VAR_GLOBAL   // PLC tag table "SDC_Carrier_TagTable"
   "Carrier_01_Carrier_In_Zone" AT %QW400 : Word;
   "Carrier_01_Carrier_Number_Echo" AT %QW402 : Word;
   "Carrier_01_Carrier_Position_Echo" AT %QD404 : DWord;
   "Carrier_01_Next_Carrier_Number" AT %QW408 : Word;
   "Carrier_01_Next_Stop_Position" AT %QD410 : DWord;
   "Carrier_01_Drive_Command_Speed" AT %QW414 : Word;
   "Carrier_01_Duplicate_Carrier_Number" AT %QW416 : Word;
   "Carrier_01_First_Duplicate_Carrier_Position" AT %QD418 : DWord;
   "Carrier_01_Second_Duplicate_Carrier_Position" AT %QD422 : DWord;
   "Carrier_01_CommandWord" AT %QW426 : Word;
   "Carrier_01_Heartbeat" AT %Q426.0 : Bool;
   "Carrier_01_Drive_Forward_Command" AT %Q426.1 : Bool;
   "Carrier_01_Fault_Reset" AT %Q426.2 : Bool;
   "Carrier_01_At_Command_Position" AT %Q426.3 : Bool;
   "Carrier_01_Duplicate_Carrier_Fault" AT %Q426.4 : Bool;
   "Carrier_01_Motion_On_Fault" AT %Q426.5 : Bool;
   "Carrier_01_Motion_Off_Fault" AT %Q426.6 : Bool;
   "Carrier_01_Carrier_Spacing_Fault" AT %Q426.7 : Bool;
   "Carrier_02_Carrier_In_Zone" AT %QW450 : Word;
   "Carrier_02_Carrier_Number_Echo" AT %QW452 : Word;
   "Carrier_02_Carrier_Position_Echo" AT %QD454 : DWord;
   "Carrier_02_Next_Carrier_Number" AT %QW458 : Word;
   "Carrier_02_Next_Stop_Position" AT %QD460 : DWord;
   "Carrier_02_Drive_Command_Speed" AT %QW464 : Word;
   "Carrier_02_Duplicate_Carrier_Number" AT %QW466 : Word;
   "Carrier_02_First_Duplicate_Carrier_Position" AT %QD468 : DWord;
   "Carrier_02_Second_Duplicate_Carrier_Position" AT %QD472 : DWord;
   "Carrier_02_CommandWord" AT %QW476 : Word;
   "Carrier_02_Heartbeat" AT %Q476.0 : Bool;
   "Carrier_02_Drive_Forward_Command" AT %Q476.1 : Bool;
   "Carrier_02_Fault_Reset" AT %Q476.2 : Bool;
   "Carrier_02_At_Command_Position" AT %Q476.3 : Bool;
   "Carrier_02_Duplicate_Carrier_Fault" AT %Q476.4 : Bool;
   "Carrier_02_Motion_On_Fault" AT %Q476.5 : Bool;
   "Carrier_02_Motion_Off_Fault" AT %Q476.6 : Bool;
   "Carrier_02_Carrier_Spacing_Fault" AT %Q476.7 : Bool;
   "Carrier_03_Carrier_In_Zone" AT %QW500 : Word;
   "Carrier_03_Carrier_Number_Echo" AT %QW502 : Word;
   "Carrier_03_Carrier_Position_Echo" AT %QD504 : DWord;
   "Carrier_03_Next_Carrier_Number" AT %QW508 : Word;
   "Carrier_03_Next_Stop_Position" AT %QD510 : DWord;
   "Carrier_03_Drive_Command_Speed" AT %QW514 : Word;
   "Carrier_03_Duplicate_Carrier_Number" AT %QW516 : Word;
   "Carrier_03_First_Duplicate_Carrier_Position" AT %QD518 : DWord;
   "Carrier_03_Second_Duplicate_Carrier_Position" AT %QD522 : DWord;
   "Carrier_03_CommandWord" AT %QW526 : Word;
   "Carrier_03_Heartbeat" AT %Q526.0 : Bool;
   "Carrier_03_Drive_Forward_Command" AT %Q526.1 : Bool;
   "Carrier_03_Fault_Reset" AT %Q526.2 : Bool;
   "Carrier_03_At_Command_Position" AT %Q526.3 : Bool;
   "Carrier_03_Duplicate_Carrier_Fault" AT %Q526.4 : Bool;
   "Carrier_03_Motion_On_Fault" AT %Q526.5 : Bool;
   "Carrier_03_Motion_Off_Fault" AT %Q526.6 : Bool;
   "Carrier_03_Carrier_Spacing_Fault" AT %Q526.7 : Bool;
   "Carrier_04_Carrier_In_Zone" AT %QW550 : Word;
   "Carrier_04_Carrier_Number_Echo" AT %QW552 : Word;
   "Carrier_04_Carrier_Position_Echo" AT %QD554 : DWord;
   "Carrier_04_Next_Carrier_Number" AT %QW558 : Word;
   "Carrier_04_Next_Stop_Position" AT %QD560 : DWord;
   "Carrier_04_Drive_Command_Speed" AT %QW564 : Word;
   "Carrier_04_Duplicate_Carrier_Number" AT %QW566 : Word;
   "Carrier_04_First_Duplicate_Carrier_Position" AT %QD568 : DWord;
   "Carrier_04_Second_Duplicate_Carrier_Position" AT %QD572 : DWord;
   "Carrier_04_CommandWord" AT %QW576 : Word;
   "Carrier_04_Heartbeat" AT %Q576.0 : Bool;
   "Carrier_04_Drive_Forward_Command" AT %Q576.1 : Bool;
   "Carrier_04_Fault_Reset" AT %Q576.2 : Bool;
   "Carrier_04_At_Command_Position" AT %Q576.3 : Bool;
   "Carrier_04_Duplicate_Carrier_Fault" AT %Q576.4 : Bool;
   "Carrier_04_Motion_On_Fault" AT %Q576.5 : Bool;
   "Carrier_04_Motion_Off_Fault" AT %Q576.6 : Bool;
   "Carrier_04_Carrier_Spacing_Fault" AT %Q576.7 : Bool;
   "Carrier_05_Carrier_In_Zone" AT %QW600 : Word;
   "Carrier_05_Carrier_Number_Echo" AT %QW602 : Word;
   "Carrier_05_Carrier_Position_Echo" AT %QD604 : DWord;
   "Carrier_05_Next_Carrier_Number" AT %QW608 : Word;
   "Carrier_05_Next_Stop_Position" AT %QD610 : DWord;
   "Carrier_05_Drive_Command_Speed" AT %QW614 : Word;
   "Carrier_05_Duplicate_Carrier_Number" AT %QW616 : Word;
   "Carrier_05_First_Duplicate_Carrier_Position" AT %QD618 : DWord;
   "Carrier_05_Second_Duplicate_Carrier_Position" AT %QD622 : DWord;
   "Carrier_05_CommandWord" AT %QW626 : Word;
   "Carrier_05_Heartbeat" AT %Q626.0 : Bool;
   "Carrier_05_Drive_Forward_Command" AT %Q626.1 : Bool;
   "Carrier_05_Fault_Reset" AT %Q626.2 : Bool;
   "Carrier_05_At_Command_Position" AT %Q626.3 : Bool;
   "Carrier_05_Duplicate_Carrier_Fault" AT %Q626.4 : Bool;
   "Carrier_05_Motion_On_Fault" AT %Q626.5 : Bool;
   "Carrier_05_Motion_Off_Fault" AT %Q626.6 : Bool;
   "Carrier_05_Carrier_Spacing_Fault" AT %Q626.7 : Bool;
   "Carrier_06_Carrier_In_Zone" AT %QW650 : Word;
   "Carrier_06_Carrier_Number_Echo" AT %QW652 : Word;
   "Carrier_06_Carrier_Position_Echo" AT %QD654 : DWord;
   "Carrier_06_Next_Carrier_Number" AT %QW658 : Word;
   "Carrier_06_Next_Stop_Position" AT %QD660 : DWord;
   "Carrier_06_Drive_Command_Speed" AT %QW664 : Word;
   "Carrier_06_Duplicate_Carrier_Number" AT %QW666 : Word;
   "Carrier_06_First_Duplicate_Carrier_Position" AT %QD668 : DWord;
   "Carrier_06_Second_Duplicate_Carrier_Position" AT %QD672 : DWord;
   "Carrier_06_CommandWord" AT %QW676 : Word;
   "Carrier_06_Heartbeat" AT %Q676.0 : Bool;
   "Carrier_06_Drive_Forward_Command" AT %Q676.1 : Bool;
   "Carrier_06_Fault_Reset" AT %Q676.2 : Bool;
   "Carrier_06_At_Command_Position" AT %Q676.3 : Bool;
   "Carrier_06_Duplicate_Carrier_Fault" AT %Q676.4 : Bool;
   "Carrier_06_Motion_On_Fault" AT %Q676.5 : Bool;
   "Carrier_06_Motion_Off_Fault" AT %Q676.6 : Bool;
   "Carrier_06_Carrier_Spacing_Fault" AT %Q676.7 : Bool;
   "Carrier_07_Carrier_In_Zone" AT %QW700 : Word;
   "Carrier_07_Carrier_Number_Echo" AT %QW702 : Word;
   "Carrier_07_Carrier_Position_Echo" AT %QD704 : DWord;
   "Carrier_07_Next_Carrier_Number" AT %QW708 : Word;
   "Carrier_07_Next_Stop_Position" AT %QD710 : DWord;
   "Carrier_07_Drive_Command_Speed" AT %QW714 : Word;
   "Carrier_07_Duplicate_Carrier_Number" AT %QW716 : Word;
   "Carrier_07_First_Duplicate_Carrier_Position" AT %QD718 : DWord;
   "Carrier_07_Second_Duplicate_Carrier_Position" AT %QD722 : DWord;
   "Carrier_07_CommandWord" AT %QW726 : Word;
   "Carrier_07_Heartbeat" AT %Q726.0 : Bool;
   "Carrier_07_Drive_Forward_Command" AT %Q726.1 : Bool;
   "Carrier_07_Fault_Reset" AT %Q726.2 : Bool;
   "Carrier_07_At_Command_Position" AT %Q726.3 : Bool;
   "Carrier_07_Duplicate_Carrier_Fault" AT %Q726.4 : Bool;
   "Carrier_07_Motion_On_Fault" AT %Q726.5 : Bool;
   "Carrier_07_Motion_Off_Fault" AT %Q726.6 : Bool;
   "Carrier_07_Carrier_Spacing_Fault" AT %Q726.7 : Bool;
   "Carrier_08_Carrier_In_Zone" AT %QW750 : Word;
   "Carrier_08_Carrier_Number_Echo" AT %QW752 : Word;
   "Carrier_08_Carrier_Position_Echo" AT %QD754 : DWord;
   "Carrier_08_Next_Carrier_Number" AT %QW758 : Word;
   "Carrier_08_Next_Stop_Position" AT %QD760 : DWord;
   "Carrier_08_Drive_Command_Speed" AT %QW764 : Word;
   "Carrier_08_Duplicate_Carrier_Number" AT %QW766 : Word;
   "Carrier_08_First_Duplicate_Carrier_Position" AT %QD768 : DWord;
   "Carrier_08_Second_Duplicate_Carrier_Position" AT %QD772 : DWord;
   "Carrier_08_CommandWord" AT %QW776 : Word;
   "Carrier_08_Heartbeat" AT %Q776.0 : Bool;
   "Carrier_08_Drive_Forward_Command" AT %Q776.1 : Bool;
   "Carrier_08_Fault_Reset" AT %Q776.2 : Bool;
   "Carrier_08_At_Command_Position" AT %Q776.3 : Bool;
   "Carrier_08_Duplicate_Carrier_Fault" AT %Q776.4 : Bool;
   "Carrier_08_Motion_On_Fault" AT %Q776.5 : Bool;
   "Carrier_08_Motion_Off_Fault" AT %Q776.6 : Bool;
   "Carrier_08_Carrier_Spacing_Fault" AT %Q776.7 : Bool;
   "Carrier_09_Carrier_In_Zone" AT %QW800 : Word;
   "Carrier_09_Carrier_Number_Echo" AT %QW802 : Word;
   "Carrier_09_Carrier_Position_Echo" AT %QD804 : DWord;
   "Carrier_09_Next_Carrier_Number" AT %QW808 : Word;
   "Carrier_09_Next_Stop_Position" AT %QD810 : DWord;
   "Carrier_09_Drive_Command_Speed" AT %QW814 : Word;
   "Carrier_09_Duplicate_Carrier_Number" AT %QW816 : Word;
   "Carrier_09_First_Duplicate_Carrier_Position" AT %QD818 : DWord;
   "Carrier_09_Second_Duplicate_Carrier_Position" AT %QD822 : DWord;
   "Carrier_09_CommandWord" AT %QW826 : Word;
   "Carrier_09_Heartbeat" AT %Q826.0 : Bool;
   "Carrier_09_Drive_Forward_Command" AT %Q826.1 : Bool;
   "Carrier_09_Fault_Reset" AT %Q826.2 : Bool;
   "Carrier_09_At_Command_Position" AT %Q826.3 : Bool;
   "Carrier_09_Duplicate_Carrier_Fault" AT %Q826.4 : Bool;
   "Carrier_09_Motion_On_Fault" AT %Q826.5 : Bool;
   "Carrier_09_Motion_Off_Fault" AT %Q826.6 : Bool;
   "Carrier_09_Carrier_Spacing_Fault" AT %Q826.7 : Bool;
   "Carrier_10_Carrier_In_Zone" AT %QW850 : Word;
   "Carrier_10_Carrier_Number_Echo" AT %QW852 : Word;
   "Carrier_10_Carrier_Position_Echo" AT %QD854 : DWord;
   "Carrier_10_Next_Carrier_Number" AT %QW858 : Word;
   "Carrier_10_Next_Stop_Position" AT %QD860 : DWord;
   "Carrier_10_Drive_Command_Speed" AT %QW864 : Word;
   "Carrier_10_Duplicate_Carrier_Number" AT %QW866 : Word;
   "Carrier_10_First_Duplicate_Carrier_Position" AT %QD868 : DWord;
   "Carrier_10_Second_Duplicate_Carrier_Position" AT %QD872 : DWord;
   "Carrier_10_CommandWord" AT %QW876 : Word;
   "Carrier_10_Heartbeat" AT %Q876.0 : Bool;
   "Carrier_10_Drive_Forward_Command" AT %Q876.1 : Bool;
   "Carrier_10_Fault_Reset" AT %Q876.2 : Bool;
   "Carrier_10_At_Command_Position" AT %Q876.3 : Bool;
   "Carrier_10_Duplicate_Carrier_Fault" AT %Q876.4 : Bool;
   "Carrier_10_Motion_On_Fault" AT %Q876.5 : Bool;
   "Carrier_10_Motion_Off_Fault" AT %Q876.6 : Bool;
   "Carrier_10_Carrier_Spacing_Fault" AT %Q876.7 : Bool;
   "Carrier_11_Carrier_In_Zone" AT %QW900 : Word;
   "Carrier_11_Carrier_Number_Echo" AT %QW902 : Word;
   "Carrier_11_Carrier_Position_Echo" AT %QD904 : DWord;
   "Carrier_11_Next_Carrier_Number" AT %QW908 : Word;
   "Carrier_11_Next_Stop_Position" AT %QD910 : DWord;
   "Carrier_11_Drive_Command_Speed" AT %QW914 : Word;
   "Carrier_11_Duplicate_Carrier_Number" AT %QW916 : Word;
   "Carrier_11_First_Duplicate_Carrier_Position" AT %QD918 : DWord;
   "Carrier_11_Second_Duplicate_Carrier_Position" AT %QD922 : DWord;
   "Carrier_11_CommandWord" AT %QW926 : Word;
   "Carrier_11_Heartbeat" AT %Q926.0 : Bool;
   "Carrier_11_Drive_Forward_Command" AT %Q926.1 : Bool;
   "Carrier_11_Fault_Reset" AT %Q926.2 : Bool;
   "Carrier_11_At_Command_Position" AT %Q926.3 : Bool;
   "Carrier_11_Duplicate_Carrier_Fault" AT %Q926.4 : Bool;
   "Carrier_11_Motion_On_Fault" AT %Q926.5 : Bool;
   "Carrier_11_Motion_Off_Fault" AT %Q926.6 : Bool;
   "Carrier_11_Carrier_Spacing_Fault" AT %Q926.7 : Bool;
   "Carrier_12_Carrier_In_Zone" AT %QW950 : Word;
   "Carrier_12_Carrier_Number_Echo" AT %QW952 : Word;
   "Carrier_12_Carrier_Position_Echo" AT %QD954 : DWord;
   "Carrier_12_Next_Carrier_Number" AT %QW958 : Word;
   "Carrier_12_Next_Stop_Position" AT %QD960 : DWord;
   "Carrier_12_Drive_Command_Speed" AT %QW964 : Word;
   "Carrier_12_Duplicate_Carrier_Number" AT %QW966 : Word;
   "Carrier_12_First_Duplicate_Carrier_Position" AT %QD968 : DWord;
   "Carrier_12_Second_Duplicate_Carrier_Position" AT %QD972 : DWord;
   "Carrier_12_CommandWord" AT %QW976 : Word;
   "Carrier_12_Heartbeat" AT %Q976.0 : Bool;
   "Carrier_12_Drive_Forward_Command" AT %Q976.1 : Bool;
   "Carrier_12_Fault_Reset" AT %Q976.2 : Bool;
   "Carrier_12_At_Command_Position" AT %Q976.3 : Bool;
   "Carrier_12_Duplicate_Carrier_Fault" AT %Q976.4 : Bool;
   "Carrier_12_Motion_On_Fault" AT %Q976.5 : Bool;
   "Carrier_12_Motion_Off_Fault" AT %Q976.6 : Bool;
   "Carrier_12_Carrier_Spacing_Fault" AT %Q976.7 : Bool;
   "Carrier_13_Carrier_In_Zone" AT %QW1000 : Word;
   "Carrier_13_Carrier_Number_Echo" AT %QW1002 : Word;
   "Carrier_13_Carrier_Position_Echo" AT %QD1004 : DWord;
   "Carrier_13_Next_Carrier_Number" AT %QW1008 : Word;
   "Carrier_13_Next_Stop_Position" AT %QD1010 : DWord;
   "Carrier_13_Drive_Command_Speed" AT %QW1014 : Word;
   "Carrier_13_Duplicate_Carrier_Number" AT %QW1016 : Word;
   "Carrier_13_First_Duplicate_Carrier_Position" AT %QD1018 : DWord;
   "Carrier_13_Second_Duplicate_Carrier_Position" AT %QD1022 : DWord;
   "Carrier_13_CommandWord" AT %QW1026 : Word;
   "Carrier_13_Heartbeat" AT %Q1026.0 : Bool;
   "Carrier_13_Drive_Forward_Command" AT %Q1026.1 : Bool;
   "Carrier_13_Fault_Reset" AT %Q1026.2 : Bool;
   "Carrier_13_At_Command_Position" AT %Q1026.3 : Bool;
   "Carrier_13_Duplicate_Carrier_Fault" AT %Q1026.4 : Bool;
   "Carrier_13_Motion_On_Fault" AT %Q1026.5 : Bool;
   "Carrier_13_Motion_Off_Fault" AT %Q1026.6 : Bool;
   "Carrier_13_Carrier_Spacing_Fault" AT %Q1026.7 : Bool;
   "Carrier_14_Carrier_In_Zone" AT %QW1050 : Word;
   "Carrier_14_Carrier_Number_Echo" AT %QW1052 : Word;
   "Carrier_14_Carrier_Position_Echo" AT %QD1054 : DWord;
   "Carrier_14_Next_Carrier_Number" AT %QW1058 : Word;
   "Carrier_14_Next_Stop_Position" AT %QD1060 : DWord;
   "Carrier_14_Drive_Command_Speed" AT %QW1064 : Word;
   "Carrier_14_Duplicate_Carrier_Number" AT %QW1066 : Word;
   "Carrier_14_First_Duplicate_Carrier_Position" AT %QD1068 : DWord;
   "Carrier_14_Second_Duplicate_Carrier_Position" AT %QD1072 : DWord;
   "Carrier_14_CommandWord" AT %QW1076 : Word;
   "Carrier_14_Heartbeat" AT %Q1076.0 : Bool;
   "Carrier_14_Drive_Forward_Command" AT %Q1076.1 : Bool;
   "Carrier_14_Fault_Reset" AT %Q1076.2 : Bool;
   "Carrier_14_At_Command_Position" AT %Q1076.3 : Bool;
   "Carrier_14_Duplicate_Carrier_Fault" AT %Q1076.4 : Bool;
   "Carrier_14_Motion_On_Fault" AT %Q1076.5 : Bool;
   "Carrier_14_Motion_Off_Fault" AT %Q1076.6 : Bool;
   "Carrier_14_Carrier_Spacing_Fault" AT %Q1076.7 : Bool;
   "Carrier_15_Carrier_In_Zone" AT %QW1100 : Word;
   "Carrier_15_Carrier_Number_Echo" AT %QW1102 : Word;
   "Carrier_15_Carrier_Position_Echo" AT %QD1104 : DWord;
   "Carrier_15_Next_Carrier_Number" AT %QW1108 : Word;
   "Carrier_15_Next_Stop_Position" AT %QD1110 : DWord;
   "Carrier_15_Drive_Command_Speed" AT %QW1114 : Word;
   "Carrier_15_Duplicate_Carrier_Number" AT %QW1116 : Word;
   "Carrier_15_First_Duplicate_Carrier_Position" AT %QD1118 : DWord;
   "Carrier_15_Second_Duplicate_Carrier_Position" AT %QD1122 : DWord;
   "Carrier_15_CommandWord" AT %QW1126 : Word;
   "Carrier_15_Heartbeat" AT %Q1126.0 : Bool;
   "Carrier_15_Drive_Forward_Command" AT %Q1126.1 : Bool;
   "Carrier_15_Fault_Reset" AT %Q1126.2 : Bool;
   "Carrier_15_At_Command_Position" AT %Q1126.3 : Bool;
   "Carrier_15_Duplicate_Carrier_Fault" AT %Q1126.4 : Bool;
   "Carrier_15_Motion_On_Fault" AT %Q1126.5 : Bool;
   "Carrier_15_Motion_Off_Fault" AT %Q1126.6 : Bool;
   "Carrier_15_Carrier_Spacing_Fault" AT %Q1126.7 : Bool;
   "Carrier_16_Carrier_In_Zone" AT %QW1150 : Word;
   "Carrier_16_Carrier_Number_Echo" AT %QW1152 : Word;
   "Carrier_16_Carrier_Position_Echo" AT %QD1154 : DWord;
   "Carrier_16_Next_Carrier_Number" AT %QW1158 : Word;
   "Carrier_16_Next_Stop_Position" AT %QD1160 : DWord;
   "Carrier_16_Drive_Command_Speed" AT %QW1164 : Word;
   "Carrier_16_Duplicate_Carrier_Number" AT %QW1166 : Word;
   "Carrier_16_First_Duplicate_Carrier_Position" AT %QD1168 : DWord;
   "Carrier_16_Second_Duplicate_Carrier_Position" AT %QD1172 : DWord;
   "Carrier_16_CommandWord" AT %QW1176 : Word;
   "Carrier_16_Heartbeat" AT %Q1176.0 : Bool;
   "Carrier_16_Drive_Forward_Command" AT %Q1176.1 : Bool;
   "Carrier_16_Fault_Reset" AT %Q1176.2 : Bool;
   "Carrier_16_At_Command_Position" AT %Q1176.3 : Bool;
   "Carrier_16_Duplicate_Carrier_Fault" AT %Q1176.4 : Bool;
   "Carrier_16_Motion_On_Fault" AT %Q1176.5 : Bool;
   "Carrier_16_Motion_Off_Fault" AT %Q1176.6 : Bool;
   "Carrier_16_Carrier_Spacing_Fault" AT %Q1176.7 : Bool;
   "Carrier_17_Carrier_In_Zone" AT %QW1200 : Word;
   "Carrier_17_Carrier_Number_Echo" AT %QW1202 : Word;
   "Carrier_17_Carrier_Position_Echo" AT %QD1204 : DWord;
   "Carrier_17_Next_Carrier_Number" AT %QW1208 : Word;
   "Carrier_17_Next_Stop_Position" AT %QD1210 : DWord;
   "Carrier_17_Drive_Command_Speed" AT %QW1214 : Word;
   "Carrier_17_Duplicate_Carrier_Number" AT %QW1216 : Word;
   "Carrier_17_First_Duplicate_Carrier_Position" AT %QD1218 : DWord;
   "Carrier_17_Second_Duplicate_Carrier_Position" AT %QD1222 : DWord;
   "Carrier_17_CommandWord" AT %QW1226 : Word;
   "Carrier_17_Heartbeat" AT %Q1226.0 : Bool;
   "Carrier_17_Drive_Forward_Command" AT %Q1226.1 : Bool;
   "Carrier_17_Fault_Reset" AT %Q1226.2 : Bool;
   "Carrier_17_At_Command_Position" AT %Q1226.3 : Bool;
   "Carrier_17_Duplicate_Carrier_Fault" AT %Q1226.4 : Bool;
   "Carrier_17_Motion_On_Fault" AT %Q1226.5 : Bool;
   "Carrier_17_Motion_Off_Fault" AT %Q1226.6 : Bool;
   "Carrier_17_Carrier_Spacing_Fault" AT %Q1226.7 : Bool;
   "Carrier_18_Carrier_In_Zone" AT %QW1250 : Word;
   "Carrier_18_Carrier_Number_Echo" AT %QW1252 : Word;
   "Carrier_18_Carrier_Position_Echo" AT %QD1254 : DWord;
   "Carrier_18_Next_Carrier_Number" AT %QW1258 : Word;
   "Carrier_18_Next_Stop_Position" AT %QD1260 : DWord;
   "Carrier_18_Drive_Command_Speed" AT %QW1264 : Word;
   "Carrier_18_Duplicate_Carrier_Number" AT %QW1266 : Word;
   "Carrier_18_First_Duplicate_Carrier_Position" AT %QD1268 : DWord;
   "Carrier_18_Second_Duplicate_Carrier_Position" AT %QD1272 : DWord;
   "Carrier_18_CommandWord" AT %QW1276 : Word;
   "Carrier_18_Heartbeat" AT %Q1276.0 : Bool;
   "Carrier_18_Drive_Forward_Command" AT %Q1276.1 : Bool;
   "Carrier_18_Fault_Reset" AT %Q1276.2 : Bool;
   "Carrier_18_At_Command_Position" AT %Q1276.3 : Bool;
   "Carrier_18_Duplicate_Carrier_Fault" AT %Q1276.4 : Bool;
   "Carrier_18_Motion_On_Fault" AT %Q1276.5 : Bool;
   "Carrier_18_Motion_Off_Fault" AT %Q1276.6 : Bool;
   "Carrier_18_Carrier_Spacing_Fault" AT %Q1276.7 : Bool;
   "Carrier_19_Carrier_In_Zone" AT %QW1300 : Word;
   "Carrier_19_Carrier_Number_Echo" AT %QW1302 : Word;
   "Carrier_19_Carrier_Position_Echo" AT %QD1304 : DWord;
   "Carrier_19_Next_Carrier_Number" AT %QW1308 : Word;
   "Carrier_19_Next_Stop_Position" AT %QD1310 : DWord;
   "Carrier_19_Drive_Command_Speed" AT %QW1314 : Word;
   "Carrier_19_Duplicate_Carrier_Number" AT %QW1316 : Word;
   "Carrier_19_First_Duplicate_Carrier_Position" AT %QD1318 : DWord;
   "Carrier_19_Second_Duplicate_Carrier_Position" AT %QD1322 : DWord;
   "Carrier_19_CommandWord" AT %QW1326 : Word;
   "Carrier_19_Heartbeat" AT %Q1326.0 : Bool;
   "Carrier_19_Drive_Forward_Command" AT %Q1326.1 : Bool;
   "Carrier_19_Fault_Reset" AT %Q1326.2 : Bool;
   "Carrier_19_At_Command_Position" AT %Q1326.3 : Bool;
   "Carrier_19_Duplicate_Carrier_Fault" AT %Q1326.4 : Bool;
   "Carrier_19_Motion_On_Fault" AT %Q1326.5 : Bool;
   "Carrier_19_Motion_Off_Fault" AT %Q1326.6 : Bool;
   "Carrier_19_Carrier_Spacing_Fault" AT %Q1326.7 : Bool;
   "Carrier_20_Carrier_In_Zone" AT %QW1350 : Word;
   "Carrier_20_Carrier_Number_Echo" AT %QW1352 : Word;
   "Carrier_20_Carrier_Position_Echo" AT %QD1354 : DWord;
   "Carrier_20_Next_Carrier_Number" AT %QW1358 : Word;
   "Carrier_20_Next_Stop_Position" AT %QD1360 : DWord;
   "Carrier_20_Drive_Command_Speed" AT %QW1364 : Word;
   "Carrier_20_Duplicate_Carrier_Number" AT %QW1366 : Word;
   "Carrier_20_First_Duplicate_Carrier_Position" AT %QD1368 : DWord;
   "Carrier_20_Second_Duplicate_Carrier_Position" AT %QD1372 : DWord;
   "Carrier_20_CommandWord" AT %QW1376 : Word;
   "Carrier_20_Heartbeat" AT %Q1376.0 : Bool;
   "Carrier_20_Drive_Forward_Command" AT %Q1376.1 : Bool;
   "Carrier_20_Fault_Reset" AT %Q1376.2 : Bool;
   "Carrier_20_At_Command_Position" AT %Q1376.3 : Bool;
   "Carrier_20_Duplicate_Carrier_Fault" AT %Q1376.4 : Bool;
   "Carrier_20_Motion_On_Fault" AT %Q1376.5 : Bool;
   "Carrier_20_Motion_Off_Fault" AT %Q1376.6 : Bool;
   "Carrier_20_Carrier_Spacing_Fault" AT %Q1376.7 : Bool;
   "Carrier_21_Carrier_In_Zone" AT %QW1400 : Word;
   "Carrier_21_Carrier_Number_Echo" AT %QW1402 : Word;
   "Carrier_21_Carrier_Position_Echo" AT %QD1404 : DWord;
   "Carrier_21_Next_Carrier_Number" AT %QW1408 : Word;
   "Carrier_21_Next_Stop_Position" AT %QD1410 : DWord;
   "Carrier_21_Drive_Command_Speed" AT %QW1414 : Word;
   "Carrier_21_Duplicate_Carrier_Number" AT %QW1416 : Word;
   "Carrier_21_First_Duplicate_Carrier_Position" AT %QD1418 : DWord;
   "Carrier_21_Second_Duplicate_Carrier_Position" AT %QD1422 : DWord;
   "Carrier_21_CommandWord" AT %QW1426 : Word;
   "Carrier_21_Heartbeat" AT %Q1426.0 : Bool;
   "Carrier_21_Drive_Forward_Command" AT %Q1426.1 : Bool;
   "Carrier_21_Fault_Reset" AT %Q1426.2 : Bool;
   "Carrier_21_At_Command_Position" AT %Q1426.3 : Bool;
   "Carrier_21_Duplicate_Carrier_Fault" AT %Q1426.4 : Bool;
   "Carrier_21_Motion_On_Fault" AT %Q1426.5 : Bool;
   "Carrier_21_Motion_Off_Fault" AT %Q1426.6 : Bool;
   "Carrier_21_Carrier_Spacing_Fault" AT %Q1426.7 : Bool;
   "Carrier_22_Carrier_In_Zone" AT %QW1450 : Word;
   "Carrier_22_Carrier_Number_Echo" AT %QW1452 : Word;
   "Carrier_22_Carrier_Position_Echo" AT %QD1454 : DWord;
   "Carrier_22_Next_Carrier_Number" AT %QW1458 : Word;
   "Carrier_22_Next_Stop_Position" AT %QD1460 : DWord;
   "Carrier_22_Drive_Command_Speed" AT %QW1464 : Word;
   "Carrier_22_Duplicate_Carrier_Number" AT %QW1466 : Word;
   "Carrier_22_First_Duplicate_Carrier_Position" AT %QD1468 : DWord;
   "Carrier_22_Second_Duplicate_Carrier_Position" AT %QD1472 : DWord;
   "Carrier_22_CommandWord" AT %QW1476 : Word;
   "Carrier_22_Heartbeat" AT %Q1476.0 : Bool;
   "Carrier_22_Drive_Forward_Command" AT %Q1476.1 : Bool;
   "Carrier_22_Fault_Reset" AT %Q1476.2 : Bool;
   "Carrier_22_At_Command_Position" AT %Q1476.3 : Bool;
   "Carrier_22_Duplicate_Carrier_Fault" AT %Q1476.4 : Bool;
   "Carrier_22_Motion_On_Fault" AT %Q1476.5 : Bool;
   "Carrier_22_Motion_Off_Fault" AT %Q1476.6 : Bool;
   "Carrier_22_Carrier_Spacing_Fault" AT %Q1476.7 : Bool;
   "Carrier_23_Carrier_In_Zone" AT %QW1500 : Word;
   "Carrier_23_Carrier_Number_Echo" AT %QW1502 : Word;
   "Carrier_23_Carrier_Position_Echo" AT %QD1504 : DWord;
   "Carrier_23_Next_Carrier_Number" AT %QW1508 : Word;
   "Carrier_23_Next_Stop_Position" AT %QD1510 : DWord;
   "Carrier_23_Drive_Command_Speed" AT %QW1514 : Word;
   "Carrier_23_Duplicate_Carrier_Number" AT %QW1516 : Word;
   "Carrier_23_First_Duplicate_Carrier_Position" AT %QD1518 : DWord;
   "Carrier_23_Second_Duplicate_Carrier_Position" AT %QD1522 : DWord;
   "Carrier_23_CommandWord" AT %QW1526 : Word;
   "Carrier_23_Heartbeat" AT %Q1526.0 : Bool;
   "Carrier_23_Drive_Forward_Command" AT %Q1526.1 : Bool;
   "Carrier_23_Fault_Reset" AT %Q1526.2 : Bool;
   "Carrier_23_At_Command_Position" AT %Q1526.3 : Bool;
   "Carrier_23_Duplicate_Carrier_Fault" AT %Q1526.4 : Bool;
   "Carrier_23_Motion_On_Fault" AT %Q1526.5 : Bool;
   "Carrier_23_Motion_Off_Fault" AT %Q1526.6 : Bool;
   "Carrier_23_Carrier_Spacing_Fault" AT %Q1526.7 : Bool;
   "Carrier_24_Carrier_In_Zone" AT %QW1550 : Word;
   "Carrier_24_Carrier_Number_Echo" AT %QW1552 : Word;
   "Carrier_24_Carrier_Position_Echo" AT %QD1554 : DWord;
   "Carrier_24_Next_Carrier_Number" AT %QW1558 : Word;
   "Carrier_24_Next_Stop_Position" AT %QD1560 : DWord;
   "Carrier_24_Drive_Command_Speed" AT %QW1564 : Word;
   "Carrier_24_Duplicate_Carrier_Number" AT %QW1566 : Word;
   "Carrier_24_First_Duplicate_Carrier_Position" AT %QD1568 : DWord;
   "Carrier_24_Second_Duplicate_Carrier_Position" AT %QD1572 : DWord;
   "Carrier_24_CommandWord" AT %QW1576 : Word;
   "Carrier_24_Heartbeat" AT %Q1576.0 : Bool;
   "Carrier_24_Drive_Forward_Command" AT %Q1576.1 : Bool;
   "Carrier_24_Fault_Reset" AT %Q1576.2 : Bool;
   "Carrier_24_At_Command_Position" AT %Q1576.3 : Bool;
   "Carrier_24_Duplicate_Carrier_Fault" AT %Q1576.4 : Bool;
   "Carrier_24_Motion_On_Fault" AT %Q1576.5 : Bool;
   "Carrier_24_Motion_Off_Fault" AT %Q1576.6 : Bool;
   "Carrier_24_Carrier_Spacing_Fault" AT %Q1576.7 : Bool;
   "Carrier_25_Carrier_In_Zone" AT %QW1600 : Word;
   "Carrier_25_Carrier_Number_Echo" AT %QW1602 : Word;
   "Carrier_25_Carrier_Position_Echo" AT %QD1604 : DWord;
   "Carrier_25_Next_Carrier_Number" AT %QW1608 : Word;
   "Carrier_25_Next_Stop_Position" AT %QD1610 : DWord;
   "Carrier_25_Drive_Command_Speed" AT %QW1614 : Word;
   "Carrier_25_Duplicate_Carrier_Number" AT %QW1616 : Word;
   "Carrier_25_First_Duplicate_Carrier_Position" AT %QD1618 : DWord;
   "Carrier_25_Second_Duplicate_Carrier_Position" AT %QD1622 : DWord;
   "Carrier_25_CommandWord" AT %QW1626 : Word;
   "Carrier_25_Heartbeat" AT %Q1626.0 : Bool;
   "Carrier_25_Drive_Forward_Command" AT %Q1626.1 : Bool;
   "Carrier_25_Fault_Reset" AT %Q1626.2 : Bool;
   "Carrier_25_At_Command_Position" AT %Q1626.3 : Bool;
   "Carrier_25_Duplicate_Carrier_Fault" AT %Q1626.4 : Bool;
   "Carrier_25_Motion_On_Fault" AT %Q1626.5 : Bool;
   "Carrier_25_Motion_Off_Fault" AT %Q1626.6 : Bool;
   "Carrier_25_Carrier_Spacing_Fault" AT %Q1626.7 : Bool;
   "Carrier_26_Carrier_In_Zone" AT %QW1650 : Word;
   "Carrier_26_Carrier_Number_Echo" AT %QW1652 : Word;
   "Carrier_26_Carrier_Position_Echo" AT %QD1654 : DWord;
   "Carrier_26_Next_Carrier_Number" AT %QW1658 : Word;
   "Carrier_26_Next_Stop_Position" AT %QD1660 : DWord;
   "Carrier_26_Drive_Command_Speed" AT %QW1664 : Word;
   "Carrier_26_Duplicate_Carrier_Number" AT %QW1666 : Word;
   "Carrier_26_First_Duplicate_Carrier_Position" AT %QD1668 : DWord;
   "Carrier_26_Second_Duplicate_Carrier_Position" AT %QD1672 : DWord;
   "Carrier_26_CommandWord" AT %QW1676 : Word;
   "Carrier_26_Heartbeat" AT %Q1676.0 : Bool;
   "Carrier_26_Drive_Forward_Command" AT %Q1676.1 : Bool;
   "Carrier_26_Fault_Reset" AT %Q1676.2 : Bool;
   "Carrier_26_At_Command_Position" AT %Q1676.3 : Bool;
   "Carrier_26_Duplicate_Carrier_Fault" AT %Q1676.4 : Bool;
   "Carrier_26_Motion_On_Fault" AT %Q1676.5 : Bool;
   "Carrier_26_Motion_Off_Fault" AT %Q1676.6 : Bool;
   "Carrier_26_Carrier_Spacing_Fault" AT %Q1676.7 : Bool;
   "Carrier_27_Carrier_In_Zone" AT %QW1700 : Word;
   "Carrier_27_Carrier_Number_Echo" AT %QW1702 : Word;
   "Carrier_27_Carrier_Position_Echo" AT %QD1704 : DWord;
   "Carrier_27_Next_Carrier_Number" AT %QW1708 : Word;
   "Carrier_27_Next_Stop_Position" AT %QD1710 : DWord;
   "Carrier_27_Drive_Command_Speed" AT %QW1714 : Word;
   "Carrier_27_Duplicate_Carrier_Number" AT %QW1716 : Word;
   "Carrier_27_First_Duplicate_Carrier_Position" AT %QD1718 : DWord;
   "Carrier_27_Second_Duplicate_Carrier_Position" AT %QD1722 : DWord;
   "Carrier_27_CommandWord" AT %QW1726 : Word;
   "Carrier_27_Heartbeat" AT %Q1726.0 : Bool;
   "Carrier_27_Drive_Forward_Command" AT %Q1726.1 : Bool;
   "Carrier_27_Fault_Reset" AT %Q1726.2 : Bool;
   "Carrier_27_At_Command_Position" AT %Q1726.3 : Bool;
   "Carrier_27_Duplicate_Carrier_Fault" AT %Q1726.4 : Bool;
   "Carrier_27_Motion_On_Fault" AT %Q1726.5 : Bool;
   "Carrier_27_Motion_Off_Fault" AT %Q1726.6 : Bool;
   "Carrier_27_Carrier_Spacing_Fault" AT %Q1726.7 : Bool;
   "Carrier_28_Carrier_In_Zone" AT %QW1750 : Word;
   "Carrier_28_Carrier_Number_Echo" AT %QW1752 : Word;
   "Carrier_28_Carrier_Position_Echo" AT %QD1754 : DWord;
   "Carrier_28_Next_Carrier_Number" AT %QW1758 : Word;
   "Carrier_28_Next_Stop_Position" AT %QD1760 : DWord;
   "Carrier_28_Drive_Command_Speed" AT %QW1764 : Word;
   "Carrier_28_Duplicate_Carrier_Number" AT %QW1766 : Word;
   "Carrier_28_First_Duplicate_Carrier_Position" AT %QD1768 : DWord;
   "Carrier_28_Second_Duplicate_Carrier_Position" AT %QD1772 : DWord;
   "Carrier_28_CommandWord" AT %QW1776 : Word;
   "Carrier_28_Heartbeat" AT %Q1776.0 : Bool;
   "Carrier_28_Drive_Forward_Command" AT %Q1776.1 : Bool;
   "Carrier_28_Fault_Reset" AT %Q1776.2 : Bool;
   "Carrier_28_At_Command_Position" AT %Q1776.3 : Bool;
   "Carrier_28_Duplicate_Carrier_Fault" AT %Q1776.4 : Bool;
   "Carrier_28_Motion_On_Fault" AT %Q1776.5 : Bool;
   "Carrier_28_Motion_Off_Fault" AT %Q1776.6 : Bool;
   "Carrier_28_Carrier_Spacing_Fault" AT %Q1776.7 : Bool;
   "Carrier_29_Carrier_In_Zone" AT %QW1800 : Word;
   "Carrier_29_Carrier_Number_Echo" AT %QW1802 : Word;
   "Carrier_29_Carrier_Position_Echo" AT %QD1804 : DWord;
   "Carrier_29_Next_Carrier_Number" AT %QW1808 : Word;
   "Carrier_29_Next_Stop_Position" AT %QD1810 : DWord;
   "Carrier_29_Drive_Command_Speed" AT %QW1814 : Word;
   "Carrier_29_Duplicate_Carrier_Number" AT %QW1816 : Word;
   "Carrier_29_First_Duplicate_Carrier_Position" AT %QD1818 : DWord;
   "Carrier_29_Second_Duplicate_Carrier_Position" AT %QD1822 : DWord;
   "Carrier_29_CommandWord" AT %QW1826 : Word;
   "Carrier_29_Heartbeat" AT %Q1826.0 : Bool;
   "Carrier_29_Drive_Forward_Command" AT %Q1826.1 : Bool;
   "Carrier_29_Fault_Reset" AT %Q1826.2 : Bool;
   "Carrier_29_At_Command_Position" AT %Q1826.3 : Bool;
   "Carrier_29_Duplicate_Carrier_Fault" AT %Q1826.4 : Bool;
   "Carrier_29_Motion_On_Fault" AT %Q1826.5 : Bool;
   "Carrier_29_Motion_Off_Fault" AT %Q1826.6 : Bool;
   "Carrier_29_Carrier_Spacing_Fault" AT %Q1826.7 : Bool;
   "Carrier_30_Carrier_In_Zone" AT %QW1850 : Word;
   "Carrier_30_Carrier_Number_Echo" AT %QW1852 : Word;
   "Carrier_30_Carrier_Position_Echo" AT %QD1854 : DWord;
   "Carrier_30_Next_Carrier_Number" AT %QW1858 : Word;
   "Carrier_30_Next_Stop_Position" AT %QD1860 : DWord;
   "Carrier_30_Drive_Command_Speed" AT %QW1864 : Word;
   "Carrier_30_Duplicate_Carrier_Number" AT %QW1866 : Word;
   "Carrier_30_First_Duplicate_Carrier_Position" AT %QD1868 : DWord;
   "Carrier_30_Second_Duplicate_Carrier_Position" AT %QD1872 : DWord;
   "Carrier_30_CommandWord" AT %QW1876 : Word;
   "Carrier_30_Heartbeat" AT %Q1876.0 : Bool;
   "Carrier_30_Drive_Forward_Command" AT %Q1876.1 : Bool;
   "Carrier_30_Fault_Reset" AT %Q1876.2 : Bool;
   "Carrier_30_At_Command_Position" AT %Q1876.3 : Bool;
   "Carrier_30_Duplicate_Carrier_Fault" AT %Q1876.4 : Bool;
   "Carrier_30_Motion_On_Fault" AT %Q1876.5 : Bool;
   "Carrier_30_Motion_Off_Fault" AT %Q1876.6 : Bool;
   "Carrier_30_Carrier_Spacing_Fault" AT %Q1876.7 : Bool;
   "Carrier_31_Carrier_In_Zone" AT %QW1900 : Word;
   "Carrier_31_Carrier_Number_Echo" AT %QW1902 : Word;
   "Carrier_31_Carrier_Position_Echo" AT %QD1904 : DWord;
   "Carrier_31_Next_Carrier_Number" AT %QW1908 : Word;
   "Carrier_31_Next_Stop_Position" AT %QD1910 : DWord;
   "Carrier_31_Drive_Command_Speed" AT %QW1914 : Word;
   "Carrier_31_Duplicate_Carrier_Number" AT %QW1916 : Word;
   "Carrier_31_First_Duplicate_Carrier_Position" AT %QD1918 : DWord;
   "Carrier_31_Second_Duplicate_Carrier_Position" AT %QD1922 : DWord;
   "Carrier_31_CommandWord" AT %QW1926 : Word;
   "Carrier_31_Heartbeat" AT %Q1926.0 : Bool;
   "Carrier_31_Drive_Forward_Command" AT %Q1926.1 : Bool;
   "Carrier_31_Fault_Reset" AT %Q1926.2 : Bool;
   "Carrier_31_At_Command_Position" AT %Q1926.3 : Bool;
   "Carrier_31_Duplicate_Carrier_Fault" AT %Q1926.4 : Bool;
   "Carrier_31_Motion_On_Fault" AT %Q1926.5 : Bool;
   "Carrier_31_Motion_Off_Fault" AT %Q1926.6 : Bool;
   "Carrier_31_Carrier_Spacing_Fault" AT %Q1926.7 : Bool;
   "Carrier_32_Carrier_In_Zone" AT %QW1950 : Word;
   "Carrier_32_Carrier_Number_Echo" AT %QW1952 : Word;
   "Carrier_32_Carrier_Position_Echo" AT %QD1954 : DWord;
   "Carrier_32_Next_Carrier_Number" AT %QW1958 : Word;
   "Carrier_32_Next_Stop_Position" AT %QD1960 : DWord;
   "Carrier_32_Drive_Command_Speed" AT %QW1964 : Word;
   "Carrier_32_Duplicate_Carrier_Number" AT %QW1966 : Word;
   "Carrier_32_First_Duplicate_Carrier_Position" AT %QD1968 : DWord;
   "Carrier_32_Second_Duplicate_Carrier_Position" AT %QD1972 : DWord;
   "Carrier_32_CommandWord" AT %QW1976 : Word;
   "Carrier_32_Heartbeat" AT %Q1976.0 : Bool;
   "Carrier_32_Drive_Forward_Command" AT %Q1976.1 : Bool;
   "Carrier_32_Fault_Reset" AT %Q1976.2 : Bool;
   "Carrier_32_At_Command_Position" AT %Q1976.3 : Bool;
   "Carrier_32_Duplicate_Carrier_Fault" AT %Q1976.4 : Bool;
   "Carrier_32_Motion_On_Fault" AT %Q1976.5 : Bool;
   "Carrier_32_Motion_Off_Fault" AT %Q1976.6 : Bool;
   "Carrier_32_Carrier_Spacing_Fault" AT %Q1976.7 : Bool;
   "Carrier_33_Carrier_In_Zone" AT %QW2000 : Word;
   "Carrier_33_Carrier_Number_Echo" AT %QW2002 : Word;
   "Carrier_33_Carrier_Position_Echo" AT %QD2004 : DWord;
   "Carrier_33_Next_Carrier_Number" AT %QW2008 : Word;
   "Carrier_33_Next_Stop_Position" AT %QD2010 : DWord;
   "Carrier_33_Drive_Command_Speed" AT %QW2014 : Word;
   "Carrier_33_Duplicate_Carrier_Number" AT %QW2016 : Word;
   "Carrier_33_First_Duplicate_Carrier_Position" AT %QD2018 : DWord;
   "Carrier_33_Second_Duplicate_Carrier_Position" AT %QD2022 : DWord;
   "Carrier_33_CommandWord" AT %QW2026 : Word;
   "Carrier_33_Heartbeat" AT %Q2026.0 : Bool;
   "Carrier_33_Drive_Forward_Command" AT %Q2026.1 : Bool;
   "Carrier_33_Fault_Reset" AT %Q2026.2 : Bool;
   "Carrier_33_At_Command_Position" AT %Q2026.3 : Bool;
   "Carrier_33_Duplicate_Carrier_Fault" AT %Q2026.4 : Bool;
   "Carrier_33_Motion_On_Fault" AT %Q2026.5 : Bool;
   "Carrier_33_Motion_Off_Fault" AT %Q2026.6 : Bool;
   "Carrier_33_Carrier_Spacing_Fault" AT %Q2026.7 : Bool;